   	
      SmartTags("SDC\DB_SDC_TS_PARAMETER\_TS_Par_HMI_Byte_00") = 0 + HMI_Nr * (Laenge_Data + HMISekDaten_Offset)  - Laenge_Data - HMISekDaten_Offset + Allg_Offset	
      SmartTags("SDC\DB_SDC_TS_PARAMETER\_TS_Par_HMI_Byte_02") = 2 + HMI_Nr * (Laenge_Data + HMISekDaten_Offset)  - Laenge_Data - HMISekDaten_Offset + Allg_Offset	
      SmartTags("SDC\DB_SDC_TS_PARAMETER\_TS_Par_HMI_Byte_04") = 4 + HMI_Nr * (Laenge_Data + HMISekDaten_Offset)  - Laenge_Data - HMISekDaten_Offset + Allg_Offset	
      SmartTags("SDC\DB_SDC_TS_PARAMETER\_TS_Par_HMI_Byte_06") = 6 + HMI_Nr * (Laenge_Data + HMISekDaten_Offset)  - Laenge_Data - HMISekDaten_Offset + Allg_Offset	
      SmartTags("SDC\DB_SDC_TS_PARAMETER\_TS_Par_HMI_Byte_08") = 8 + HMI_Nr * (Laenge_Data + HMISekDaten_Offset)  - Laenge_Data - HMISekDaten_Offset + Allg_Offset	
      SmartTags("SDC\DB_SDC_TS_PARAMETER\_TS_Par_HMI_Byte_09") = 9 + HMI_Nr * (Laenge_Data + HMISekDaten_Offset)  - Laenge_Data - HMISekDaten_Offset + Allg_Offset	
      SmartTags("SDC\DB_SDC_TS_PARAMETER\_TS_Par_HMI_Byte_10") = 10 + HMI_Nr * (Laenge_Data + HMISekDaten_Offset)  - Laenge_Data - HMISekDaten_Offset + Allg_Offset	
      SmartTags("SDC\DB_SDC_TS_PARAMETER\_TS_Par_HMI_Byte_12") = 12 + HMI_Nr * (Laenge_Data + HMISekDaten_Offset)  - Laenge_Data - HMISekDaten_Offset + Allg_Offset		
      SmartTags("SDC\DB_SDC_TS_PARAMETER\_TS_Par_HMI_Byte_14") = 14 + HMI_Nr * (Laenge_Data + HMISekDaten_Offset)  - Laenge_Data - HMISekDaten_Offset + Allg_Offset	
      SmartTags("SDC\DB_SDC_TS_PARAMETER\_TS_Par_HMI_Byte_16") = 16 + HMI_Nr * (Laenge_Data + HMISekDaten_Offset)  - Laenge_Data - HMISekDaten_Offset + Allg_Offset	
      SmartTags("SDC\DB_SDC_TS_PARAMETER\_TS_Par_HMI_Byte_18") = 18 + HMI_Nr * (Laenge_Data + HMISekDaten_Offset)  - Laenge_Data - HMISekDaten_Offset + Allg_Offset	
      SmartTags("SDC\DB_SDC_TS_PARAMETER\_TS_Par_HMI_Byte_19") = 19 + HMI_Nr * (Laenge_Data + HMISekDaten_Offset)  - Laenge_Data - HMISekDaten_Offset + Allg_Offset
   
      SmartTags("SDC\DB_SDC_TS_PARAMETER\_TS_Par_Allg_Byte_00") =  0 + HMI_Nr * (Laenge_Data + HMISekDaten_Offset)  - Laenge_Data + Allg_Offset
      SmartTags("SDC\DB_SDC_TS_PARAMETER\_TS_Par_Allg_Byte_02") =  2 + HMI_Nr * (Laenge_Data + HMISekDaten_Offset)  - Laenge_Data + Allg_Offset  
      SmartTags("SDC\DB_SDC_TS_PARAMETER\_TS_Par_Allg_Byte_06") =  6 + HMI_Nr * (Laenge_Data + HMISekDaten_Offset)  - Laenge_Data + Allg_Offset  
      SmartTags("SDC\DB_SDC_TS_PARAMETER\_TS_Par_Allg_Byte_10") = 10 + HMI_Nr * (Laenge_Data + HMISekDaten_Offset)  - Laenge_Data + Allg_Offset   
      SmartTags("SDC\DB_SDC_TS_PARAMETER\_TS_Par_Allg_Byte_22") = 22 + HMI_Nr * (Laenge_Data + HMISekDaten_Offset)  - Laenge_Data + Allg_Offset   
      SmartTags("SDC\DB_SDC_TS_PARAMETER\_TS_Par_Allg_Byte_24") = 24 + HMI_Nr * (Laenge_Data + HMISekDaten_Offset)  - Laenge_Data + Allg_Offset   
      SmartTags("SDC\DB_SDC_TS_PARAMETER\_TS_Par_Allg_Byte_26") = 26 + HMI_Nr * (Laenge_Data + HMISekDaten_Offset)  - Laenge_Data + Allg_Offset 
      SmartTags("SDC\DB_SDC_TS_PARAMETER\_TS_Par_Allg_Byte_27") = 27 + HMI_Nr * (Laenge_Data + HMISekDaten_Offset)  - Laenge_Data + Allg_Offset      
      SmartTags("SDC\DB_SDC_TS_PARAMETER\_TS_Par_Allg_Byte_28") = 28 + HMI_Nr * (Laenge_Data + HMISekDaten_Offset)  - Laenge_Data + Allg_Offset  
      SmartTags("SDC\DB_SDC_TS_PARAMETER\_TS_Par_Allg_Byte_29") = 29 + HMI_Nr * (Laenge_Data + HMISekDaten_Offset)  - Laenge_Data + Allg_Offset     
      SmartTags("SDC\DB_SDC_TS_PARAMETER\_TS_Par_Allg_Byte_30") = 30 + HMI_Nr * (Laenge_Data + HMISekDaten_Offset)  - Laenge_Data + Allg_Offset  
      SmartTags("SDC\DB_SDC_TS_PARAMETER\_TS_Par_Allg_Byte_32") = 32 + HMI_Nr * (Laenge_Data + HMISekDaten_Offset)  - Laenge_Data + Allg_Offset 
      SmartTags("SDC\DB_SDC_TS_PARAMETER\_TS_Par_Allg_Byte_36") = 36 + HMI_Nr * (Laenge_Data + HMISekDaten_Offset)  - Laenge_Data + Allg_Offset 
         
      SmartTags("SDC\DB_SDC_TS_PARAMETER\_TS_Par_Profil_Byte_00") =  0 + HMI_Nr * (Laenge_Data + HMISekDaten_Offset)  - Laenge_Data + Allg_Offset + Profil_Offset + TS_Profil_Nr * Laenge_Profil - Laenge_Profil
      SmartTags("SDC\DB_SDC_TS_PARAMETER\_TS_Par_Profil_Byte_02") =  2 + HMI_Nr * (Laenge_Data + HMISekDaten_Offset)  - Laenge_Data + Allg_Offset + Profil_Offset + TS_Profil_Nr * Laenge_Profil - Laenge_Profil
      SmartTags("SDC\DB_SDC_TS_PARAMETER\_TS_Par_Profil_Byte_04") =  4 + HMI_Nr * (Laenge_Data + HMISekDaten_Offset)  - Laenge_Data + Allg_Offset + Profil_Offset + TS_Profil_Nr * Laenge_Profil - Laenge_Profil
      SmartTags("SDC\DB_SDC_TS_PARAMETER\_TS_Par_Profil_Byte_06") =  6 + HMI_Nr * (Laenge_Data + HMISekDaten_Offset)  - Laenge_Data + Allg_Offset + Profil_Offset + TS_Profil_Nr * Laenge_Profil - Laenge_Profil   	 
      SmartTags("SDC\DB_SDC_TS_PARAMETER\_TS_Par_Profil_Byte_08") =  8 + HMI_Nr * (Laenge_Data + HMISekDaten_Offset)  - Laenge_Data + Allg_Offset + Profil_Offset + TS_Profil_Nr * Laenge_Profil - Laenge_Profil
      SmartTags("SDC\DB_SDC_TS_PARAMETER\_TS_Par_Profil_Byte_10") = 10 + HMI_Nr * (Laenge_Data + HMISekDaten_Offset)  - Laenge_Data + Allg_Offset + Profil_Offset + TS_Profil_Nr * Laenge_Profil - Laenge_Profil
      SmartTags("SDC\DB_SDC_TS_PARAMETER\_TS_Par_Profil_Byte_12") = 12 + HMI_Nr * (Laenge_Data + HMISekDaten_Offset)  - Laenge_Data + Allg_Offset + Profil_Offset + TS_Profil_Nr * Laenge_Profil - Laenge_Profil
      SmartTags("SDC\DB_SDC_TS_PARAMETER\_TS_Par_Profil_Byte_14") = 14 + HMI_Nr * (Laenge_Data + HMISekDaten_Offset)  - Laenge_Data + Allg_Offset + Profil_Offset + TS_Profil_Nr * Laenge_Profil - Laenge_Profil   	  
      SmartTags("SDC\DB_SDC_TS_PARAMETER\_TS_Par_Profil_Byte_16") = 16 + HMI_Nr * (Laenge_Data + HMISekDaten_Offset)  - Laenge_Data + Allg_Offset + Profil_Offset + TS_Profil_Nr * Laenge_Profil - Laenge_Profil
      SmartTags("SDC\DB_SDC_TS_PARAMETER\_TS_Par_Profil_Byte_18") = 18 + HMI_Nr * (Laenge_Data + HMISekDaten_Offset)  - Laenge_Data + Allg_Offset + Profil_Offset + TS_Profil_Nr * Laenge_Profil - Laenge_Profil
      SmartTags("SDC\DB_SDC_TS_PARAMETER\_TS_Par_Profil_Byte_20") = 20 + HMI_Nr * (Laenge_Data + HMISekDaten_Offset)  - Laenge_Data + Allg_Offset + Profil_Offset + TS_Profil_Nr * Laenge_Profil - Laenge_Profil
      SmartTags("SDC\DB_SDC_TS_PARAMETER\_TS_Par_Profil_Byte_22") = 22 + HMI_Nr * (Laenge_Data + HMISekDaten_Offset)  - Laenge_Data + Allg_Offset + Profil_Offset + TS_Profil_Nr * Laenge_Profil - Laenge_Profil   	 
      SmartTags("SDC\DB_SDC_TS_PARAMETER\_TS_Par_Profil_Byte_24") = 24 + HMI_Nr * (Laenge_Data + HMISekDaten_Offset)  - Laenge_Data + Allg_Offset + Profil_Offset + TS_Profil_Nr * Laenge_Profil - Laenge_Profil
      SmartTags("SDC\DB_SDC_TS_PARAMETER\_TS_Par_Profil_Byte_26") = 26 + HMI_Nr * (Laenge_Data + HMISekDaten_Offset)  - Laenge_Data + Allg_Offset + Profil_Offset + TS_Profil_Nr * Laenge_Profil - Laenge_Profil
      SmartTags("SDC\DB_SDC_TS_PARAMETER\_TS_Par_Profil_Byte_28") = 28 + HMI_Nr * (Laenge_Data + HMISekDaten_Offset)  - Laenge_Data + Allg_Offset + Profil_Offset + TS_Profil_Nr * Laenge_Profil - Laenge_Profil
      SmartTags("SDC\DB_SDC_TS_PARAMETER\_TS_Par_Profil_Byte_30") = 30 + HMI_Nr * (Laenge_Data + HMISekDaten_Offset)  - Laenge_Data + Allg_Offset + Profil_Offset + TS_Profil_Nr * Laenge_Profil - Laenge_Profil   	
      SmartTags("SDC\DB_SDC_TS_PARAMETER\_TS_Par_Profil_Byte_32") = 32 + HMI_Nr * (Laenge_Data + HMISekDaten_Offset)  - Laenge_Data + Allg_Offset + Profil_Offset + TS_Profil_Nr * Laenge_Profil - Laenge_Profil
      SmartTags("SDC\DB_SDC_TS_PARAMETER\_TS_Par_Profil_Byte_34") = 34 + HMI_Nr * (Laenge_Data + HMISekDaten_Offset)  - Laenge_Data + Allg_Offset + Profil_Offset + TS_Profil_Nr * Laenge_Profil - Laenge_Profil
      SmartTags("SDC\DB_SDC_TS_PARAMETER\_TS_Par_Profil_Byte_36") = 36 + HMI_Nr * (Laenge_Data + HMISekDaten_Offset)  - Laenge_Data + Allg_Offset + Profil_Offset + TS_Profil_Nr * Laenge_Profil - Laenge_Profil   	 
      SmartTags("SDC\DB_SDC_TS_PARAMETER\_TS_Par_Profil_Byte_38") = 38 + HMI_Nr * (Laenge_Data + HMISekDaten_Offset)  - Laenge_Data + Allg_Offset + Profil_Offset + TS_Profil_Nr * Laenge_Profil - Laenge_Profil
      SmartTags("SDC\DB_SDC_TS_PARAMETER\_TS_Par_Profil_Byte_40") = 40 + HMI_Nr * (Laenge_Data + HMISekDaten_Offset)  - Laenge_Data + Allg_Offset + Profil_Offset + TS_Profil_Nr * Laenge_Profil - Laenge_Profil
      SmartTags("SDC\DB_SDC_TS_PARAMETER\_TS_Par_Profil_Byte_42") = 42 + HMI_Nr * (Laenge_Data + HMISekDaten_Offset)  - Laenge_Data + Allg_Offset + Profil_Offset + TS_Profil_Nr * Laenge_Profil - Laenge_Profil
   
      SmartTags("SDC\DB_SDC_TS_PARAMETER\_TS_Par_Profil+1_Byte_00") =  0 + HMI_Nr * (Laenge_Data + HMISekDaten_Offset)  - Laenge_Data + Allg_Offset + Profil_Offset + (TS_Profil_Nr +1) * Laenge_Profil - Laenge_Profil
      SmartTags("SDC\DB_SDC_TS_PARAMETER\_TS_Par_Profil+1_Byte_02") =  2 + HMI_Nr * (Laenge_Data + HMISekDaten_Offset)  - Laenge_Data + Allg_Offset + Profil_Offset + (TS_Profil_Nr +1) * Laenge_Profil - Laenge_Profil
      SmartTags("SDC\DB_SDC_TS_PARAMETER\_TS_Par_Profil+1_Byte_04") =  4 + HMI_Nr * (Laenge_Data + HMISekDaten_Offset)  - Laenge_Data + Allg_Offset + Profil_Offset + (TS_Profil_Nr +1) * Laenge_Profil - Laenge_Profil
      SmartTags("SDC\DB_SDC_TS_PARAMETER\_TS_Par_Profil+1_Byte_06") =  6 + HMI_Nr * (Laenge_Data + HMISekDaten_Offset)  - Laenge_Data + Allg_Offset + Profil_Offset + (TS_Profil_Nr +1) * Laenge_Profil - Laenge_Profil   	 
      SmartTags("SDC\DB_SDC_TS_PARAMETER\_TS_Par_Profil+1_Byte_08") =  8 + HMI_Nr * (Laenge_Data + HMISekDaten_Offset)  - Laenge_Data + Allg_Offset + Profil_Offset + (TS_Profil_Nr +1) * Laenge_Profil - Laenge_Profil
      SmartTags("SDC\DB_SDC_TS_PARAMETER\_TS_Par_Profil+1_Byte_10") = 10 + HMI_Nr * (Laenge_Data + HMISekDaten_Offset)  - Laenge_Data + Allg_Offset + Profil_Offset + (TS_Profil_Nr +1) * Laenge_Profil - Laenge_Profil
      SmartTags("SDC\DB_SDC_TS_PARAMETER\_TS_Par_Profil+1_Byte_12") = 12 + HMI_Nr * (Laenge_Data + HMISekDaten_Offset)  - Laenge_Data + Allg_Offset + Profil_Offset + (TS_Profil_Nr +1) * Laenge_Profil - Laenge_Profil
      SmartTags("SDC\DB_SDC_TS_PARAMETER\_TS_Par_Profil+1_Byte_14") = 14 + HMI_Nr * (Laenge_Data + HMISekDaten_Offset)  - Laenge_Data + Allg_Offset + Profil_Offset + (TS_Profil_Nr +1) * Laenge_Profil - Laenge_Profil   	  
      SmartTags("SDC\DB_SDC_TS_PARAMETER\_TS_Par_Profil+1_Byte_16") = 16 + HMI_Nr * (Laenge_Data + HMISekDaten_Offset)  - Laenge_Data + Allg_Offset + Profil_Offset + (TS_Profil_Nr +1) * Laenge_Profil - Laenge_Profil
      SmartTags("SDC\DB_SDC_TS_PARAMETER\_TS_Par_Profil+1_Byte_18") = 18 + HMI_Nr * (Laenge_Data + HMISekDaten_Offset)  - Laenge_Data + Allg_Offset + Profil_Offset + (TS_Profil_Nr +1) * Laenge_Profil - Laenge_Profil
      SmartTags("SDC\DB_SDC_TS_PARAMETER\_TS_Par_Profil+1_Byte_20") = 20 + HMI_Nr * (Laenge_Data + HMISekDaten_Offset)  - Laenge_Data + Allg_Offset + Profil_Offset + (TS_Profil_Nr +1) * Laenge_Profil - Laenge_Profil
      SmartTags("SDC\DB_SDC_TS_PARAMETER\_TS_Par_Profil+1_Byte_22") = 22 + HMI_Nr * (Laenge_Data + HMISekDaten_Offset)  - Laenge_Data + Allg_Offset + Profil_Offset + (TS_Profil_Nr +1) * Laenge_Profil - Laenge_Profil   	 
      SmartTags("SDC\DB_SDC_TS_PARAMETER\_TS_Par_Profil+1_Byte_24") = 24 + HMI_Nr * (Laenge_Data + HMISekDaten_Offset)  - Laenge_Data + Allg_Offset + Profil_Offset + (TS_Profil_Nr +1) * Laenge_Profil - Laenge_Profil
      SmartTags("SDC\DB_SDC_TS_PARAMETER\_TS_Par_Profil+1_Byte_26") = 26 + HMI_Nr * (Laenge_Data + HMISekDaten_Offset)  - Laenge_Data + Allg_Offset + Profil_Offset + (TS_Profil_Nr +1) * Laenge_Profil - Laenge_Profil
      SmartTags("SDC\DB_SDC_TS_PARAMETER\_TS_Par_Profil+1_Byte_28") = 28 + HMI_Nr * (Laenge_Data + HMISekDaten_Offset)  - Laenge_Data + Allg_Offset + Profil_Offset + (TS_Profil_Nr +1) * Laenge_Profil - Laenge_Profil
      SmartTags("SDC\DB_SDC_TS_PARAMETER\_TS_Par_Profil+1_Byte_30") = 30 + HMI_Nr * (Laenge_Data + HMISekDaten_Offset)  - Laenge_Data + Allg_Offset + Profil_Offset + (TS_Profil_Nr +1) * Laenge_Profil - Laenge_Profil   	
      SmartTags("SDC\DB_SDC_TS_PARAMETER\_TS_Par_Profil+1_Byte_32") = 32 + HMI_Nr * (Laenge_Data + HMISekDaten_Offset)  - Laenge_Data + Allg_Offset + Profil_Offset + (TS_Profil_Nr +1) * Laenge_Profil - Laenge_Profil
      SmartTags("SDC\DB_SDC_TS_PARAMETER\_TS_Par_Profil+1_Byte_34") = 34 + HMI_Nr * (Laenge_Data + HMISekDaten_Offset)  - Laenge_Data + Allg_Offset + Profil_Offset + (TS_Profil_Nr +1) * Laenge_Profil - Laenge_Profil
      SmartTags("SDC\DB_SDC_TS_PARAMETER\_TS_Par_Profil+1_Byte_36") = 36 + HMI_Nr * (Laenge_Data + HMISekDaten_Offset)  - Laenge_Data + Allg_Offset + Profil_Offset + (TS_Profil_Nr +1) * Laenge_Profil - Laenge_Profil   	 
      SmartTags("SDC\DB_SDC_TS_PARAMETER\_TS_Par_Profil+1_Byte_38") = 38 + HMI_Nr * (Laenge_Data + HMISekDaten_Offset)  - Laenge_Data + Allg_Offset + Profil_Offset + (TS_Profil_Nr +1) * Laenge_Profil - Laenge_Profil
      SmartTags("SDC\DB_SDC_TS_PARAMETER\_TS_Par_Profil+1_Byte_40") = 40 + HMI_Nr * (Laenge_Data + HMISekDaten_Offset)  - Laenge_Data + Allg_Offset + Profil_Offset + (TS_Profil_Nr +1) * Laenge_Profil - Laenge_Profil
      SmartTags("SDC\DB_SDC_TS_PARAMETER\_TS_Par_Profil+1_Byte_42") = 42 + HMI_Nr * (Laenge_Data + HMISekDaten_Offset)  - Laenge_Data + Allg_Offset + Profil_Offset + (TS_Profil_Nr +1) * Laenge_Profil - Laenge_Profil
   
      SmartTags("SDC\DB_SDC_TS_PARAMETER\DB_SDC_TS_PARAMETER_HMI.HMI[XX].PROFIL_Nr") = TS_Profil_Nr
      SmartTags("SDC\DB_SDC_TS_PARAMETER\DB_SDC_TS_PARAMETER_HMI.HMI[XX].SEK_Nr") = TS_Nr
   
   '##############################################
   ' VISU Sucht sich Sektions daten:
   '##############################################
   'TS_Profil_Nr = SmartTags("SDC\DB_SDC_TS_PARAMETER\_TS_Profil_Nr")
   'TS_Nr = SmartTags("SDC\DB_SDC_TS_PARAMETER\_TS_Nr")
   'Laenge_Data = SmartTags("SDC\DB_SDC_TS_PARAMETER\DB_SDC_TS_PARAMETER_1.HEADER.LAENGE_SEK_DATA")
   'Laenge_Profil = SmartTags("SDC\DB_SDC_TS_PARAMETER\DB_SDC_TS_PARAMETER_1.HEADER.LAENGE_PROFIL_DATA")
   'Allg_Offset = SmartTags("SDC\DB_SDC_TS_PARAMETER\DB_SDC_TS_PARAMETER_1.HEADER.START_DAT")
   'Profil_Offset = SmartTags("SDC\DB_SDC_TS_PARAMETER\DB_SDC_TS_PARAMETER_1.HEADER.OFFEST_PROFIL")
   
   ' search for DB Number / DBB Number --------------------------------------------
   'If SmartTags("SDC\DB_SDC_TS_PARAMETER\_TS_Nr") >= SmartTags("SDC\DB_SDC_TS_PARAMETER\DB_SDC_TS_PARAMETER_1.HEADER.MIN_NR_SEK") And SmartTags("SDC\DB_SDC_TS_PARAMETER\_TS_Nr") <= SmartTags("SDC\DB_SDC_TS_PARAMETER\DB_SDC_TS_PARAMETER_1.HEADER.MAX_NR_SEK") Then
    
   '   SmartTags("SDC\DB_SDC_TS_PARAMETER\_TS_DB_Nr") = SmartTags("SDC\DB_SDC_TS_PARAMETER\DB_SDC_TS_PARAMETER_1.HEADER.DB_NR")   
   
   '   SmartTags("SDC\DB_SDC_TS_PARAMETER\_TS_Par_Allg_Byte_00") =  0 + TS_Nr * Laenge_Data - Laenge_Data + Allg_Offset
   '   SmartTags("SDC\DB_SDC_TS_PARAMETER\_TS_Par_Allg_Byte_02") =  2 + TS_Nr * Laenge_Data - Laenge_Data + Allg_Offset  
   '   SmartTags("SDC\DB_SDC_TS_PARAMETER\_TS_Par_Allg_Byte_06") =  6 + TS_Nr * Laenge_Data - Laenge_Data + Allg_Offset  
   '   SmartTags("SDC\DB_SDC_TS_PARAMETER\_TS_Par_Allg_Byte_10") = 10 + TS_Nr * Laenge_Data - Laenge_Data + Allg_Offset   
   '   SmartTags("SDC\DB_SDC_TS_PARAMETER\_TS_Par_Allg_Byte_22") = 22 + TS_Nr * Laenge_Data - Laenge_Data + Allg_Offset   
   '   SmartTags("SDC\DB_SDC_TS_PARAMETER\_TS_Par_Allg_Byte_24") = 24 + TS_Nr * Laenge_Data - Laenge_Data + Allg_Offset   
   '   SmartTags("SDC\DB_SDC_TS_PARAMETER\_TS_Par_Allg_Byte_26") = 26 + TS_Nr * Laenge_Data - Laenge_Data + Allg_Offset 
   '   SmartTags("SDC\DB_SDC_TS_PARAMETER\_TS_Par_Allg_Byte_27") = 27 + TS_Nr * Laenge_Data - Laenge_Data + Allg_Offset      
   '   SmartTags("SDC\DB_SDC_TS_PARAMETER\_TS_Par_Allg_Byte_28") = 28 + TS_Nr * Laenge_Data - Laenge_Data + Allg_Offset  
   '   SmartTags("SDC\DB_SDC_TS_PARAMETER\_TS_Par_Allg_Byte_29") = 29 + TS_Nr * Laenge_Data - Laenge_Data + Allg_Offset     
   '   SmartTags("SDC\DB_SDC_TS_PARAMETER\_TS_Par_Allg_Byte_30") = 30 + TS_Nr * Laenge_Data - Laenge_Data + Allg_Offset  
   '   SmartTags("SDC\DB_SDC_TS_PARAMETER\_TS_Par_Allg_Byte_32") = 32 + TS_Nr * Laenge_Data - Laenge_Data + Allg_Offset 
   '   SmartTags("SDC\DB_SDC_TS_PARAMETER\_TS_Par_Allg_Byte_36") = 36 + TS_Nr * Laenge_Data - Laenge_Data + Allg_Offset 
         
   '   SmartTags("SDC\DB_SDC_TS_PARAMETER\_TS_Par_Profil_Byte_00") =  0 + TS_Nr * Laenge_Data - Laenge_Data + Allg_Offset + Profil_Offset + TS_Profil_Nr * Laenge_Profil - Laenge_Profil
   '   SmartTags("SDC\DB_SDC_TS_PARAMETER\_TS_Par_Profil_Byte_02") =  2 + TS_Nr * Laenge_Data - Laenge_Data + Allg_Offset + Profil_Offset + TS_Profil_Nr * Laenge_Profil - Laenge_Profil
   '   SmartTags("SDC\DB_SDC_TS_PARAMETER\_TS_Par_Profil_Byte_04") =  4 + TS_Nr * Laenge_Data - Laenge_Data + Allg_Offset + Profil_Offset + TS_Profil_Nr * Laenge_Profil - Laenge_Profil
   '   SmartTags("SDC\DB_SDC_TS_PARAMETER\_TS_Par_Profil_Byte_06") =  6 + TS_Nr * Laenge_Data - Laenge_Data + Allg_Offset + Profil_Offset + TS_Profil_Nr * Laenge_Profil - Laenge_Profil   	 
   '   SmartTags("SDC\DB_SDC_TS_PARAMETER\_TS_Par_Profil_Byte_08") =  8 + TS_Nr * Laenge_Data - Laenge_Data + Allg_Offset + Profil_Offset + TS_Profil_Nr * Laenge_Profil - Laenge_Profil
   '   SmartTags("SDC\DB_SDC_TS_PARAMETER\_TS_Par_Profil_Byte_10") = 10 + TS_Nr * Laenge_Data - Laenge_Data + Allg_Offset + Profil_Offset + TS_Profil_Nr * Laenge_Profil - Laenge_Profil
   '   SmartTags("SDC\DB_SDC_TS_PARAMETER\_TS_Par_Profil_Byte_12") = 12 + TS_Nr * Laenge_Data - Laenge_Data + Allg_Offset + Profil_Offset + TS_Profil_Nr * Laenge_Profil - Laenge_Profil
   '   SmartTags("SDC\DB_SDC_TS_PARAMETER\_TS_Par_Profil_Byte_14") = 14 + TS_Nr * Laenge_Data - Laenge_Data + Allg_Offset + Profil_Offset + TS_Profil_Nr * Laenge_Profil - Laenge_Profil   	  
   '   SmartTags("SDC\DB_SDC_TS_PARAMETER\_TS_Par_Profil_Byte_16") = 16 + TS_Nr * Laenge_Data - Laenge_Data + Allg_Offset + Profil_Offset + TS_Profil_Nr * Laenge_Profil - Laenge_Profil
   '   SmartTags("SDC\DB_SDC_TS_PARAMETER\_TS_Par_Profil_Byte_18") = 18 + TS_Nr * Laenge_Data - Laenge_Data + Allg_Offset + Profil_Offset + TS_Profil_Nr * Laenge_Profil - Laenge_Profil
   '   SmartTags("SDC\DB_SDC_TS_PARAMETER\_TS_Par_Profil_Byte_20") = 20 + TS_Nr * Laenge_Data - Laenge_Data + Allg_Offset + Profil_Offset + TS_Profil_Nr * Laenge_Profil - Laenge_Profil
   '   SmartTags("SDC\DB_SDC_TS_PARAMETER\_TS_Par_Profil_Byte_22") = 22 + TS_Nr * Laenge_Data - Laenge_Data + Allg_Offset + Profil_Offset + TS_Profil_Nr * Laenge_Profil - Laenge_Profil   	 
   '   SmartTags("SDC\DB_SDC_TS_PARAMETER\_TS_Par_Profil_Byte_24") = 24 + TS_Nr * Laenge_Data - Laenge_Data + Allg_Offset + Profil_Offset + TS_Profil_Nr * Laenge_Profil - Laenge_Profil
   '   SmartTags("SDC\DB_SDC_TS_PARAMETER\_TS_Par_Profil_Byte_26") = 26 + TS_Nr * Laenge_Data - Laenge_Data + Allg_Offset + Profil_Offset + TS_Profil_Nr * Laenge_Profil - Laenge_Profil
   '   SmartTags("SDC\DB_SDC_TS_PARAMETER\_TS_Par_Profil_Byte_28") = 28 + TS_Nr * Laenge_Data - Laenge_Data + Allg_Offset + Profil_Offset + TS_Profil_Nr * Laenge_Profil - Laenge_Profil
   '   SmartTags("SDC\DB_SDC_TS_PARAMETER\_TS_Par_Profil_Byte_30") = 30 + TS_Nr * Laenge_Data - Laenge_Data + Allg_Offset + Profil_Offset + TS_Profil_Nr * Laenge_Profil - Laenge_Profil   	
   '   SmartTags("SDC\DB_SDC_TS_PARAMETER\_TS_Par_Profil_Byte_32") = 32 + TS_Nr * Laenge_Data - Laenge_Data + Allg_Offset + Profil_Offset + TS_Profil_Nr * Laenge_Profil - Laenge_Profil
   '   SmartTags("SDC\DB_SDC_TS_PARAMETER\_TS_Par_Profil_Byte_34") = 34 + TS_Nr * Laenge_Data - Laenge_Data + Allg_Offset + Profil_Offset + TS_Profil_Nr * Laenge_Profil - Laenge_Profil
   '   SmartTags("SDC\DB_SDC_TS_PARAMETER\_TS_Par_Profil_Byte_36") = 36 + TS_Nr * Laenge_Data - Laenge_Data + Allg_Offset + Profil_Offset + TS_Profil_Nr * Laenge_Profil - Laenge_Profil   	 
   '   SmartTags("SDC\DB_SDC_TS_PARAMETER\_TS_Par_Profil_Byte_38") = 38 + TS_Nr * Laenge_Data - Laenge_Data + Allg_Offset + Profil_Offset + TS_Profil_Nr * Laenge_Profil - Laenge_Profil
   '   SmartTags("SDC\DB_SDC_TS_PARAMETER\_TS_Par_Profil_Byte_40") = 40 + TS_Nr * Laenge_Data - Laenge_Data + Allg_Offset + Profil_Offset + TS_Profil_Nr * Laenge_Profil - Laenge_Profil
   '   SmartTags("SDC\DB_SDC_TS_PARAMETER\_TS_Par_Profil_Byte_42") = 42 + TS_Nr * Laenge_Data - Laenge_Data + Allg_Offset + Profil_Offset + TS_Profil_Nr * Laenge_Profil - Laenge_Profil
   
   'End If
   
   'If SmartTags("SDC\DB_SDC_TS_PARAMETER\_TS_Nr") >= SmartTags("SDC\DB_SDC_TS_PARAMETER\DB_SDC_TS_PARAMETER_2.HEADER.MIN_NR_SEK") And SmartTags("SDC\DB_SDC_TS_PARAMETER\_TS_Nr") <= SmartTags("SDC\DB_SDC_TS_PARAMETER\DB_SDC_TS_PARAMETER_2.HEADER.MAX_NR_SEK") Then
   
   '  SmartTags("SDC\DB_SDC_TS_PARAMETER\_TS_DB_Nr") = SmartTags("SDC\DB_SDC_TS_PARAMETER\DB_SDC_TS_PARAMETER_2.HEADER.DB_NR")   
   
   '   TS_Nr = TS_Nr - SmartTags("SDC\DB_SDC_TS_PARAMETER\DB_SDC_TS_PARAMETER_2.HEADER.MIN_NR_SEK") + 1
   
   '  SmartTags("SDC\DB_SDC_TS_PARAMETER\_TS_Par_Allg_Byte_00") =  0 + TS_Nr * Laenge_Data - Laenge_Data + Allg_Offset
   '   SmartTags("SDC\DB_SDC_TS_PARAMETER\_TS_Par_Allg_Byte_02") =  2 + TS_Nr * Laenge_Data - Laenge_Data + Allg_Offset  
   '   SmartTags("SDC\DB_SDC_TS_PARAMETER\_TS_Par_Allg_Byte_06") =  6 + TS_Nr * Laenge_Data - Laenge_Data + Allg_Offset  
   '   SmartTags("SDC\DB_SDC_TS_PARAMETER\_TS_Par_Allg_Byte_10") = 10 + TS_Nr * Laenge_Data - Laenge_Data + Allg_Offset   
   '   SmartTags("SDC\DB_SDC_TS_PARAMETER\_TS_Par_Allg_Byte_22") = 22 + TS_Nr * Laenge_Data - Laenge_Data + Allg_Offset   
   '   SmartTags("SDC\DB_SDC_TS_PARAMETER\_TS_Par_Allg_Byte_24") = 24 + TS_Nr * Laenge_Data - Laenge_Data + Allg_Offset   
   '   SmartTags("SDC\DB_SDC_TS_PARAMETER\_TS_Par_Allg_Byte_26") = 26 + TS_Nr * Laenge_Data - Laenge_Data + Allg_Offset 
   '   SmartTags("SDC\DB_SDC_TS_PARAMETER\_TS_Par_Allg_Byte_27") = 27 + TS_Nr * Laenge_Data - Laenge_Data + Allg_Offset      
   '   SmartTags("SDC\DB_SDC_TS_PARAMETER\_TS_Par_Allg_Byte_28") = 28 + TS_Nr * Laenge_Data - Laenge_Data + Allg_Offset  
   '   SmartTags("SDC\DB_SDC_TS_PARAMETER\_TS_Par_Allg_Byte_29") = 29 + TS_Nr * Laenge_Data - Laenge_Data + Allg_Offset     
   '   SmartTags("SDC\DB_SDC_TS_PARAMETER\_TS_Par_Allg_Byte_30") = 30 + TS_Nr * Laenge_Data - Laenge_Data + Allg_Offset  
   '   SmartTags("SDC\DB_SDC_TS_PARAMETER\_TS_Par_Allg_Byte_32") = 32 + TS_Nr * Laenge_Data - Laenge_Data + Allg_Offset 
   '   SmartTags("SDC\DB_SDC_TS_PARAMETER\_TS_Par_Allg_Byte_36") = 36 + TS_Nr * Laenge_Data - Laenge_Data + Allg_Offset 
         
   '   SmartTags("SDC\DB_SDC_TS_PARAMETER\_TS_Par_Profil_Byte_00") =  0 + TS_Nr * Laenge_Data - Laenge_Data + Allg_Offset + Profil_Offset + TS_Profil_Nr * Laenge_Profil - Laenge_Profil
   '   SmartTags("SDC\DB_SDC_TS_PARAMETER\_TS_Par_Profil_Byte_02") =  2 + TS_Nr * Laenge_Data - Laenge_Data + Allg_Offset + Profil_Offset + TS_Profil_Nr * Laenge_Profil - Laenge_Profil
   '   SmartTags("SDC\DB_SDC_TS_PARAMETER\_TS_Par_Profil_Byte_04") =  4 + TS_Nr * Laenge_Data - Laenge_Data + Allg_Offset + Profil_Offset + TS_Profil_Nr * Laenge_Profil - Laenge_Profil
   '   SmartTags("SDC\DB_SDC_TS_PARAMETER\_TS_Par_Profil_Byte_06") =  6 + TS_Nr * Laenge_Data - Laenge_Data + Allg_Offset + Profil_Offset + TS_Profil_Nr * Laenge_Profil - Laenge_Profil   	 
   '   SmartTags("SDC\DB_SDC_TS_PARAMETER\_TS_Par_Profil_Byte_08") =  8 + TS_Nr * Laenge_Data - Laenge_Data + Allg_Offset + Profil_Offset + TS_Profil_Nr * Laenge_Profil - Laenge_Profil
   '   SmartTags("SDC\DB_SDC_TS_PARAMETER\_TS_Par_Profil_Byte_10") = 10 + TS_Nr * Laenge_Data - Laenge_Data + Allg_Offset + Profil_Offset + TS_Profil_Nr * Laenge_Profil - Laenge_Profil
   '   SmartTags("SDC\DB_SDC_TS_PARAMETER\_TS_Par_Profil_Byte_12") = 12 + TS_Nr * Laenge_Data - Laenge_Data + Allg_Offset + Profil_Offset + TS_Profil_Nr * Laenge_Profil - Laenge_Profil
   '   SmartTags("SDC\DB_SDC_TS_PARAMETER\_TS_Par_Profil_Byte_14") = 14 + TS_Nr * Laenge_Data - Laenge_Data + Allg_Offset + Profil_Offset + TS_Profil_Nr * Laenge_Profil - Laenge_Profil   	  
   '   SmartTags("SDC\DB_SDC_TS_PARAMETER\_TS_Par_Profil_Byte_16") = 16 + TS_Nr * Laenge_Data - Laenge_Data + Allg_Offset + Profil_Offset + TS_Profil_Nr * Laenge_Profil - Laenge_Profil
   '   SmartTags("SDC\DB_SDC_TS_PARAMETER\_TS_Par_Profil_Byte_18") = 18 + TS_Nr * Laenge_Data - Laenge_Data + Allg_Offset + Profil_Offset + TS_Profil_Nr * Laenge_Profil - Laenge_Profil
   '   SmartTags("SDC\DB_SDC_TS_PARAMETER\_TS_Par_Profil_Byte_20") = 20 + TS_Nr * Laenge_Data - Laenge_Data + Allg_Offset + Profil_Offset + TS_Profil_Nr * Laenge_Profil - Laenge_Profil
   '   SmartTags("SDC\DB_SDC_TS_PARAMETER\_TS_Par_Profil_Byte_22") = 22 + TS_Nr * Laenge_Data - Laenge_Data + Allg_Offset + Profil_Offset + TS_Profil_Nr * Laenge_Profil - Laenge_Profil   	 
   '   SmartTags("SDC\DB_SDC_TS_PARAMETER\_TS_Par_Profil_Byte_24") = 24 + TS_Nr * Laenge_Data - Laenge_Data + Allg_Offset + Profil_Offset + TS_Profil_Nr * Laenge_Profil - Laenge_Profil
   '   SmartTags("SDC\DB_SDC_TS_PARAMETER\_TS_Par_Profil_Byte_26") = 26 + TS_Nr * Laenge_Data - Laenge_Data + Allg_Offset + Profil_Offset + TS_Profil_Nr * Laenge_Profil - Laenge_Profil
   '   SmartTags("SDC\DB_SDC_TS_PARAMETER\_TS_Par_Profil_Byte_28") = 28 + TS_Nr * Laenge_Data - Laenge_Data + Allg_Offset + Profil_Offset + TS_Profil_Nr * Laenge_Profil - Laenge_Profil
   '   SmartTags("SDC\DB_SDC_TS_PARAMETER\_TS_Par_Profil_Byte_30") = 30 + TS_Nr * Laenge_Data - Laenge_Data + Allg_Offset + Profil_Offset + TS_Profil_Nr * Laenge_Profil - Laenge_Profil   	
   '   SmartTags("SDC\DB_SDC_TS_PARAMETER\_TS_Par_Profil_Byte_32") = 32 + TS_Nr * Laenge_Data - Laenge_Data + Allg_Offset + Profil_Offset + TS_Profil_Nr * Laenge_Profil - Laenge_Profil
   '   SmartTags("SDC\DB_SDC_TS_PARAMETER\_TS_Par_Profil_Byte_34") = 34 + TS_Nr * Laenge_Data - Laenge_Data + Allg_Offset + Profil_Offset + TS_Profil_Nr * Laenge_Profil - Laenge_Profil
   '   SmartTags("SDC\DB_SDC_TS_PARAMETER\_TS_Par_Profil_Byte_36") = 36 + TS_Nr * Laenge_Data - Laenge_Data + Allg_Offset + Profil_Offset + TS_Profil_Nr * Laenge_Profil - Laenge_Profil   	 
   '   SmartTags("SDC\DB_SDC_TS_PARAMETER\_TS_Par_Profil_Byte_38") = 38 + TS_Nr * Laenge_Data - Laenge_Data + Allg_Offset + Profil_Offset + TS_Profil_Nr * Laenge_Profil - Laenge_Profil
   '   SmartTags("SDC\DB_SDC_TS_PARAMETER\_TS_Par_Profil_Byte_40") = 40 + TS_Nr * Laenge_Data - Laenge_Data + Allg_Offset + Profil_Offset + TS_Profil_Nr * Laenge_Profil - Laenge_Profil
   '   SmartTags("SDC\DB_SDC_TS_PARAMETER\_TS_Par_Profil_Byte_42") = 42 + TS_Nr * Laenge_Data - Laenge_Data + Allg_Offset + Profil_Offset + TS_Profil_Nr * Laenge_Profil - Laenge_Profil
   
   'End If

VB script "SDC_TS_REFERENCE"
   'HINWEIS:
   ' Beim Erstellen von Skripten können Sie mit <Strg+Leertaste> vordefinierte 
   ' Systemfunktionen in das neue Skript einbinden.
   ' Das HMIRuntime-Objekt ermöglicht einfachen Zugriff auf die Objekte des
   ' WinCC flexible Objektmodells, ihre Methoden und ihre Eigenschaften.
   ' Für ein komfortables Auswählen einer Objektreferenz betätigen Sie bitte <Alt+Rechts>.
   ' Komplexe Skripte können Sie mit Sprachelementen der Programmiersprache
   ' VBScript erstellen.
   ' Der Zugriff auf WinCC flexible Variablen erfolgt direkt über den Variablennamen,
   ' z.B. Tag = 5
   
   '________________________________________________________________________________
   '
   
   ' Groiß Andreas
   ' Siemens AG Österreich 
   ' Linz Kraußstraße 1-7 
   ' RC-AT I-IA AS-FA-SO-AE2
   ' 02.08.2013
   
   Dim TS_Nr ' Sektion Number
   Dim Laenge_Data ' Länge TS REFERENCE
   Dim Allg_Offset ' Allg REFERENCE Offset
   
   ' INIT-------------------------------------------------------------
   SmartTags("SDC\DB_SDC_TS_REFERENCE\_TS_Ref_DB_Nr") = SmartTags("DB_SDC_TS_REFERENCE_1_HEADER.DB_NR")
   
   SmartTags("SDC\DB_SDC_TS_REFERENCE\_TS_Ref_Nr") = TS_Nr_IN
   
   If (SmartTags("SDC\DB_SDC_TS_REFERENCE\_TS_Ref_Nr") < SmartTags("DB_SDC_GLOBAL_SEK_MIN")) Or (SmartTags("SDC\DB_SDC_TS_REFERENCE\_TS_Ref_Nr") > SmartTags("DB_SDC_GLOBAL_SEK_MAX")) Then
   	SmartTags("SDC\DB_SDC_TS_REFERENCE\_TS_Ref_Nr") = 	SmartTags("DB_SDC_GLOBAL_SEK_MIN")
   End If	
   
   If (SmartTags("SDC\DB_SDC_TS_REFERENCE\_TS_Ref_Nr") < 1) Then
   	SmartTags("SDC\DB_SDC_TS_REFERENCE\_TS_Ref_Nr") = 1
   End If	
   
   
   TS_Nr = SmartTags("SDC\DB_SDC_TS_REFERENCE\_TS_Ref_Nr")
   Laenge_Data = SmartTags("DB_SDC_TS_REFERENCE_1_HEADER.LAENGE_SEK_DATA")
   Allg_Offset = SmartTags("DB_SDC_TS_REFERENCE_1_HEADER.START_DAT")
   
   ' search for DB Number / DBB Number --------------------------------------------
   If SmartTags("SDC\DB_SDC_TS_REFERENCE\_TS_Ref_Nr") >= SmartTags("DB_SDC_TS_REFERENCE_1_HEADER.MIN_NR_SEK") And SmartTags("SDC\DB_SDC_TS_REFERENCE\_TS_Ref_Nr") <= SmartTags("DB_SDC_TS_REFERENCE_1_HEADER.MAX_NR_SEK") Then
    
      SmartTags("SDC\DB_SDC_TS_REFERENCE\_TS_Ref_DB_Nr") = SmartTags("DB_SDC_TS_REFERENCE_1_HEADER.DB_NR")   
   
      SmartTags("SDC\DB_SDC_TS_REFERENCE\_TS_Ref_Byte_00")  =   0 + TS_Nr * Laenge_Data - Laenge_Data + Allg_Offset
      SmartTags("SDC\DB_SDC_TS_REFERENCE\_TS_Ref_Byte_16")  =  16 + TS_Nr * Laenge_Data - Laenge_Data + Allg_Offset  
      SmartTags("SDC\DB_SDC_TS_REFERENCE\_TS_Ref_Byte_32")  =  32 + TS_Nr * Laenge_Data - Laenge_Data + Allg_Offset  
      SmartTags("SDC\DB_SDC_TS_REFERENCE\_TS_Ref_Byte_48")  =  48 + TS_Nr * Laenge_Data - Laenge_Data + Allg_Offset   
      SmartTags("SDC\DB_SDC_TS_REFERENCE\_TS_Ref_Byte_64")  =  64 + TS_Nr * Laenge_Data - Laenge_Data + Allg_Offset   
      SmartTags("SDC\DB_SDC_TS_REFERENCE\_TS_Ref_Byte_80")  =  80 + TS_Nr * Laenge_Data - Laenge_Data + Allg_Offset   
      SmartTags("SDC\DB_SDC_TS_REFERENCE\_TS_Ref_Byte_96")  =  96 + TS_Nr * Laenge_Data - Laenge_Data + Allg_Offset 
      SmartTags("SDC\DB_SDC_TS_REFERENCE\_TS_Ref_Byte_112") = 112 + TS_Nr * Laenge_Data - Laenge_Data + Allg_Offset      
    
   End If
   
   If SmartTags("SDC\DB_SDC_TS_REFERENCE\_TS_Ref_Nr") >= SmartTags("DB_SDC_TS_REFERENCE_2_HEADER.MIN_NR_SEK") And SmartTags("SDC\DB_SDC_TS_REFERENCE\_TS_Ref_Nr") <= SmartTags("DB_SDC_TS_REFERENCE_2_HEADER.MAX_NR_SEK") Then
   
      SmartTags("SDC\DB_SDC_TS_REFERENCE\_TS_Ref_DB_Nr") = SmartTags("DB_SDC_TS_REFERENCE_2_HEADER.DB_NR")   
   
      TS_Nr = TS_Nr - SmartTags("DB_SDC_TS_REFERENCE_2_HEADER.MIN_NR_SEK") + 1
   
      SmartTags("SDC\DB_SDC_TS_REFERENCE\_TS_Ref_Byte_00")  =   0 + TS_Nr * Laenge_Data - Laenge_Data + Allg_Offset
      SmartTags("SDC\DB_SDC_TS_REFERENCE\_TS_Ref_Byte_16")  =  16 + TS_Nr * Laenge_Data - Laenge_Data + Allg_Offset  
      SmartTags("SDC\DB_SDC_TS_REFERENCE\_TS_Ref_Byte_32")  =  32 + TS_Nr * Laenge_Data - Laenge_Data + Allg_Offset  
      SmartTags("SDC\DB_SDC_TS_REFERENCE\_TS_Ref_Byte_48")  =  48 + TS_Nr * Laenge_Data - Laenge_Data + Allg_Offset   
      SmartTags("SDC\DB_SDC_TS_REFERENCE\_TS_Ref_Byte_64")  =  64 + TS_Nr * Laenge_Data - Laenge_Data + Allg_Offset   
      SmartTags("SDC\DB_SDC_TS_REFERENCE\_TS_Ref_Byte_80")  =  80 + TS_Nr * Laenge_Data - Laenge_Data + Allg_Offset   
      SmartTags("SDC\DB_SDC_TS_REFERENCE\_TS_Ref_Byte_96")  =  96 + TS_Nr * Laenge_Data - Laenge_Data + Allg_Offset 
      SmartTags("SDC\DB_SDC_TS_REFERENCE\_TS_Ref_Byte_112") = 112 + TS_Nr * Laenge_Data - Laenge_Data + Allg_Offset      
    
   End If
   
   If SmartTags("SDC\DB_SDC_TS_REFERENCE\_TS_Ref_Nr") >= SmartTags("DB_SDC_TS_REFERENCE_3_HEADER.MIN_NR_SEK") And SmartTags("SDC\DB_SDC_TS_REFERENCE\_TS_Ref_Nr") <= SmartTags("DB_SDC_TS_REFERENCE_3_HEADER.MAX_NR_SEK") Then
   
      SmartTags("SDC\DB_SDC_TS_REFERENCE\_TS_Ref_DB_Nr") = SmartTags("DB_SDC_TS_REFERENCE_3_HEADER.DB_NR")   
   
      TS_Nr = TS_Nr - SmartTags("DB_SDC_TS_REFERENCE_3_HEADER.MIN_NR_SEK") + 1
   
      SmartTags("SDC\DB_SDC_TS_REFERENCE\_TS_Ref_Byte_00")  =   0 + TS_Nr * Laenge_Data - Laenge_Data + Allg_Offset
      SmartTags("SDC\DB_SDC_TS_REFERENCE\_TS_Ref_Byte_16")  =  16 + TS_Nr * Laenge_Data - Laenge_Data + Allg_Offset  
      SmartTags("SDC\DB_SDC_TS_REFERENCE\_TS_Ref_Byte_32")  =  32 + TS_Nr * Laenge_Data - Laenge_Data + Allg_Offset  
      SmartTags("SDC\DB_SDC_TS_REFERENCE\_TS_Ref_Byte_48")  =  48 + TS_Nr * Laenge_Data - Laenge_Data + Allg_Offset   
      SmartTags("SDC\DB_SDC_TS_REFERENCE\_TS_Ref_Byte_64")  =  64 + TS_Nr * Laenge_Data - Laenge_Data + Allg_Offset   
      SmartTags("SDC\DB_SDC_TS_REFERENCE\_TS_Ref_Byte_80")  =  80 + TS_Nr * Laenge_Data - Laenge_Data + Allg_Offset   
      SmartTags("SDC\DB_SDC_TS_REFERENCE\_TS_Ref_Byte_96")  =  96 + TS_Nr * Laenge_Data - Laenge_Data + Allg_Offset 
      SmartTags("SDC\DB_SDC_TS_REFERENCE\_TS_Ref_Byte_112") = 112 + TS_Nr * Laenge_Data - Laenge_Data + Allg_Offset      
    
   End If
   
   If SmartTags("SDC\DB_SDC_TS_REFERENCE\_TS_Ref_Nr") >= SmartTags("DB_SDC_TS_REFERENCE_4_HEADER.MIN_NR_SEK") And SmartTags("SDC\DB_SDC_TS_REFERENCE\_TS_Ref_Nr") <= SmartTags("DB_SDC_TS_REFERENCE_4_HEADER.MAX_NR_SEK") Then
   
      SmartTags("SDC\DB_SDC_TS_REFERENCE\_TS_Ref_DB_Nr") = SmartTags("DB_SDC_TS_REFERENCE_4_HEADER.DB_NR")   
   
      TS_Nr = TS_Nr - SmartTags("DB_SDC_TS_REFERENCE_4_HEADER.MIN_NR_SEK") + 1
   
      SmartTags("SDC\DB_SDC_TS_REFERENCE\_TS_Ref_Byte_00")  =   0 + TS_Nr * Laenge_Data - Laenge_Data + Allg_Offset
      SmartTags("SDC\DB_SDC_TS_REFERENCE\_TS_Ref_Byte_16")  =  16 + TS_Nr * Laenge_Data - Laenge_Data + Allg_Offset  
      SmartTags("SDC\DB_SDC_TS_REFERENCE\_TS_Ref_Byte_32")  =  32 + TS_Nr * Laenge_Data - Laenge_Data + Allg_Offset  
      SmartTags("SDC\DB_SDC_TS_REFERENCE\_TS_Ref_Byte_48")  =  48 + TS_Nr * Laenge_Data - Laenge_Data + Allg_Offset   
      SmartTags("SDC\DB_SDC_TS_REFERENCE\_TS_Ref_Byte_64")  =  64 + TS_Nr * Laenge_Data - Laenge_Data + Allg_Offset   
      SmartTags("SDC\DB_SDC_TS_REFERENCE\_TS_Ref_Byte_80")  =  80 + TS_Nr * Laenge_Data - Laenge_Data + Allg_Offset   
      SmartTags("SDC\DB_SDC_TS_REFERENCE\_TS_Ref_Byte_96")  =  96 + TS_Nr * Laenge_Data - Laenge_Data + Allg_Offset 
      SmartTags("SDC\DB_SDC_TS_REFERENCE\_TS_Ref_Byte_112") = 112 + TS_Nr * Laenge_Data - Laenge_Data + Allg_Offset      
    
   End If
   
